// TIA Portal project "FORMING_1500_PLC" (V15)

(* hardware
DEVICE "1.Forming_Machine_PN"  KTP1200 Basic PN
   slot 0: "1.Forming_Machine_PN"  KTP1200 Basic PN  6AV2 123-2MB03-0AX0  15.0.0.0
   slot 1: "HMI_RT_1"  KTP1200 Basic PN  6AV2 123-2MB03-0AX0  15.0.0.0
   slot 5: "Forming_Machine.IE_CP_1"  PROFINET Interface  15.0.0.0
      slot 1: "PROFINET Interface_1"  PROFINET Interface
         slot 1: "Port_1"  Port
DEVICE "GSD device_2"  GSD.Device
   slot 0: "Rack_0"  Rail
DEVICE "GSD device_8"  GSD.Device
   slot 0: "Rack_0"  Rail
DEVICE "GSD device_5"  GSD.Device
   slot 0: "Rack_0"  Rail
DEVICE "GSD device_6"  GSD.Device
   slot 0: "Rack_0"  Rail
DEVICE "GSD device_7"  GSD.Device
   slot 0: "Rack_0"  Rail
DEVICE "GSD device_9"  GSD.Device
   slot 0: "Rack_0"  Rail
DEVICE "GSD device_4"  GSD.Device
   slot 0: "Rack_0"  Rail
DEVICE "GSD device_3"  GSD.Device
   slot 0: "Rack_0"  Rail
DEVICE "GSD device_11"  GSD.Device
   slot 0: "Rack_0"  Rail
DEVICE "GSD device_12"  GSD.Device
   slot 0: "Rack_0"  Rail
DEVICE "GSD device_13"  GSD.Device
   slot 0: "Rack_0"  Rail
DEVICE "GSD device_14"  GSD.Device
   slot 0: "Rack_0"  Rail
DEVICE "GSD device_10"  GSD.Device
   slot 0: "Rack_0"  Rail
DEVICE "GSD device_16"  GSD.Device
   slot 0: "Rack_0"  Rail
DEVICE "GSD device_17"  GSD.Device
   slot 0: "Rack_0"  Rail
DEVICE "GSD device_18"  GSD.Device
   slot 0: "Rack_0"  Rail
DEVICE "GSD device_19"  GSD.Device
   slot 0: "Rack_0"  Rail
DEVICE "GSD device_20"  GSD.Device
   slot 0: "Rack_0"  Rail
DEVICE "GSD device_15"  GSD.Device
   slot 0: "Rack_0"  Rail
DEVICE "GSD device_21"  GSD.Device
   slot 0: "Rack_0"  Rail
DEVICE "GSD device_22"  GSD.Device
   slot 0: "Rack_0"  Rail
DEVICE "GSD device_23"  GSD.Device
   slot 0: "Rack_0"  Rail
DEVICE "S71500/ET200MP station_2"  S7-1500 station
   slot 0: "Rail_0"  Rack  6ES7 590-1***0-0AA0
   slot 0: "PM 190W 120/230VAC"  PM 190W 120/230VAC  6EP1333-4BA00
   slot 1: "FORMING LINE 7 PLC_1"  CPU 1511-1 PN  6ES7 511-1AK02-0AB0  V2.5
      slot 3: "CPU display_1"  6ES7591-1AA00-0AA0
   slot 2: "CM 1542-5_1"  CM 1542-5  6GK7 542-5DX00-0XE0  V2.0
   slot 3: "DI 32x24VDC BA_3"  DI 32x24VDC BA  6ES7 521-1BL10-0AA0  V1.0
   slot 4: "DQ 16x24VDC/0.5A BA_1"  DQ 16x24VDC/0.5A BA  6ES7 522-1BH10-0AA0  V1.0
   slot 5: "DI 32x24VDC BA_1"  DI 32x24VDC BA  6ES7 521-1BL10-0AA0  V1.0
   slot 6: "DI 32x24VDC BA_2"  DI 32x24VDC BA  6ES7 521-1BL10-0AA0  V1.0
*)

// ===== PLC "FORMING LINE 7 PLC_1"  CPU 1511-1 PN =====

VAR_GLOBAL   // PLC tag table "Default tag table"
   "PHOTOCELL OF KIBBLER" AT %I7.4 : Bool;
   "KIBBLER 1 CMD" AT %M28.0 : Bool;
   "KIBBLER CLCKWISE / ANTI CLCKWISE 2" AT %Q124.2 : Bool;
   "KIBBLER 2 CMD" AT %M28.1 : Bool;
   "DELAY KIBBLER 1" AT %T14 : Timer;
   "KIBBLER CLCKWISE / ANTI CLCKWISE 1" AT %Q124.1 : Bool;
   "DELAY KIBBLER 1 RESET" AT %T15 : Timer;
   "DELAY KIBBLER 2" AT %T16 : Timer;
   "DELAY KIBBLER 2 RESET" AT %T17 : Timer;
   "INPUT METAL DETECT ALARM" AT %I7.5 : Bool;
   "input metal detect cmd a" AT %M60.1 : Bool;
   "TIMER RESET ALARM OUT METAL DETECT" AT %T9 : Timer;
   "TIMER INPUT METAL DETECT ALARM" AT %T25 : Timer;
   "input metal detect cmd b" AT %M60.0 : Bool;
   "trigger_alarm_metal_detect" AT %M38.3 : Bool;
   "ALARM OUTPUT WHEN METAL DETECT" AT %Q124.4 : Bool;
   "trigger_time_lap_metal_detect" AT %M38.4 : Bool;
   "TIME LAP WHEN METAL DETECTED" AT %Q124.0 : Bool;
   "RESET TIME LAP WHEN METAL DETECT" AT %T23 : Timer;
   "trigger_sync_addres_13" AT %M31.6 : Bool;
   "trigger_sync_addres_17 a" AT %M32.2 : Bool;
   "trigger_sync_addres_3" AT %M30.4 : Bool;
   "trigger_sync_addres_4" AT %M30.5 : Bool;
   "trigger_sync_addres_5" AT %M30.6 : Bool;
   "trigger_sync_addres_6" AT %M30.7 : Bool;
   "trigger_sync_addres_7" AT %M31.0 : Bool;
   "trigger_sync_addres_8" AT %M31.1 : Bool;
   "trigger_sync_addres_9" AT %M31.2 : Bool;
   "trigger_sync_addres_10" AT %M31.3 : Bool;
   "trigger_sync_addres_11" AT %M31.4 : Bool;
   "trigger_sync_addres_12" AT %M31.5 : Bool;
   "trigger_sync_addres_14" AT %M31.7 : Bool;
   "trigger_sync_addres_15" AT %M32.0 : Bool;
   "trigger_sync_addres_16" AT %M32.1 : Bool;
   "trigger_sync_addres_17 b" AT %M33.2 : Bool;
   "trigger_sync_addres_19" AT %M32.4 : Bool;
   "trigger_sync_addres_21" AT %M32.6 : Bool;
   "trigger_sync_addres_22" AT %M32.7 : Bool;
   "trigger_sync_addres_23" AT %M33.0 : Bool;
   "SB1" AT %I125.0 : Bool;
   "SB2" AT %I125.1 : Bool;
   "SB3" AT %I125.2 : Bool;
   "SB4" AT %I125.3 : Bool;
   "SB5" AT %I125.4 : Bool;
   "SB6" AT %I125.5 : Bool;
   "SB7" AT %I125.6 : Bool;
   "SB8" AT %I125.7 : Bool;
   "SB9" AT %I6.0 : Bool;
   "SB10" AT %I6.1 : Bool;
   "SB11" AT %I6.2 : Bool;
   "SB12" AT %I6.3 : Bool;
   "SB13" AT %I6.4 : Bool;
   "profibus addres 2 fault" AT %M90.1 : Bool;
   "profibus addres 3 fault" AT %M90.2 : Bool;
   "profibus addres 4 fault" AT %M90.3 : Bool;
   "profibus addres 5 fault" AT %M90.4 : Bool;
   "profibus addres 6 fault" AT %M90.5 : Bool;
   "profibus addres 7 fault" AT %M90.6 : Bool;
   "profibus addres 8 fault" AT %M90.7 : Bool;
   "profibus addres 9 fault" AT %M91.0 : Bool;
   "profibus addres 10 fault" AT %M91.1 : Bool;
   "profibus addres 11 fault" AT %M91.2 : Bool;
   "profibus addres 12 fault" AT %M91.3 : Bool;
   "profibus addres 13 fault" AT %M91.4 : Bool;
   "profibus addres 14 fault" AT %M91.5 : Bool;
   "profibus addres 15 fault" AT %M91.6 : Bool;
   "profibus addres 16 fault" AT %M91.7 : Bool;
   "profibus addres 17 fault" AT %M92.0 : Bool;
   "profibus addres 18 fault" AT %M92.1 : Bool;
   "profibus addres 19 fault" AT %M92.2 : Bool;
   "profibus addres 20 fault" AT %M92.3 : Bool;
   "profibus addres 21 fault" AT %M92.4 : Bool;
   "profibus addres 22 fault" AT %M92.5 : Bool;
   "profibus addres 23 fault" AT %M92.6 : Bool;
   "delay10ms_2" AT %T11 : Timer;
   "delay10ms_1" AT %T10 : Timer;
   "delay10ms_4" AT %T13 : Timer;
   "delay10ms_3" AT %T12 : Timer;
   "ROTARY MOULDER MODE" AT %I7.0 : Bool;
   "ROTARY CUTTER MODE" AT %I7.1 : Bool;
   "EMERGENCY" AT %I7.6 : Bool;
   "EMC PRESSED" AT %M92.7 : Bool;
END_VAR

VAR_GLOBAL   // PLC tag table "STEP7 classic symbols"
   "DECREASE_ADDRS_3" AT %I0.5 : Bool;
   "DECREASE_ADDRS_2" AT %I0.3 : Bool;
   "DECREASE_ADDRS_23" AT %I5.5 : Bool;
   "DECREASE_ADDRS_22" AT %I5.3 : Bool;
   "DECREASE_ADDRS_21" AT %I5.1 : Bool;
   "DECREASE_ADDRS_20" AT %I4.7 : Bool;
   "DECREASE_ADDRS_19" AT %I4.5 : Bool;
   "DECREASE_ADDRS_18" AT %I4.3 : Bool;
   "DECREASE_ADDRS_17" AT %I4.1 : Bool;
   "DECREASE_ADDRS_16" AT %I3.7 : Bool;
   "DECREASE_ADDRS_15" AT %I3.5 : Bool;
   "DECREASE_ADDRS_14" AT %I3.3 : Bool;
   "DECREASE_ADDRS_13" AT %I3.1 : Bool;
   "DECREASE_ADDRS_12" AT %I2.7 : Bool;
   "DECREASE_ADDRS_11" AT %I2.5 : Bool;
   "P_MAV_PROFIBUS_23" AT %IW510 : Word;
   "P_CTW_PROFIBUS_7" AT %QW316 : Word;
   "P_CTW_PROFIBUS_6" AT %QW304 : Word;
   "P_CTW_PROFIBUS_5" AT %QW292 : Word;
   "P_CTW_PROFIBUS_4" AT %QW280 : Word;
   "P_CTW_PROFIBUS_3" AT %QW268 : Word;
   "P_CTW_PROFIBUS_2" AT %QW256 : Word;
   "P_CTW_PROFIBUS_11" AT %QW364 : Word;
   "P_CTW_PROFIBUS_10" AT %QW352 : Word;
   "P_CTW_PROFIBUS_9" AT %QW340 : Word;
   "P_CTW_PROFIBUS_8" AT %QW328 : Word;
   "P_CTW_PROFIBUS_13" AT %QW388 : Word;
   "P_CTW_PROFIBUS_12" AT %QW376 : Word;
   "P_CTW_PROFIBUS_15" AT %QW412 : Word;
   "P_CTW_PROFIBUS_14" AT %QW400 : Word;
   "INCREASE_CMD_7" AT %M10.5 : Bool;
   "INCREASE_CMD_6" AT %M10.4 : Bool;
   "INCREASE_CMD_5" AT %M10.3 : Bool;
   "INCREASE_CMD_4" AT %M10.2 : Bool;
   "INCREASE_CMD_3" AT %M10.1 : Bool;
   "INCREASE_CMD_2" AT %M10.0 : Bool;
   "INCREASE_CMD_23" AT %M12.5 : Bool;
   "INCREASE_CMD_22" AT %M12.4 : Bool;
   "INCREASE_CMD_21" AT %M12.3 : Bool;
   "INCREASE_CMD_20" AT %M12.2 : Bool;
   "INCREASE_CMD_19" AT %M12.1 : Bool;
   "INCREASE_CMD_18" AT %M12.0 : Bool;
   "INCREASE_CMD_17" AT %M11.7 : Bool;
   "INCREASE_CMD_16" AT %M11.6 : Bool;
   "INCREASE_CMD_15" AT %M11.5 : Bool;
   "P_MRV_PROFIBUS_8" AT %QW330 : Word;
   "P_MRV_PROFIBUS_7" AT %QW318 : Word;
   "P_MRV_PROFIBUS_12" AT %QW378 : Word;
   "P_MRV_PROFIBUS_11" AT %QW366 : Word;
   "P_MRV_PROFIBUS_10" AT %QW354 : Word;
   "P_MRV_PROFIBUS_15" AT %QW414 : Word;
   "P_MRV_PROFIBUS_14" AT %QW402 : Word;
   "P_MRV_PROFIBUS_13" AT %QW390 : Word;
   "P_MRV_PROFIBUS_18" AT %QW450 : Word;
   "P_MRV_PROFIBUS_17" AT %QW438 : Word;
   "P_MRV_PROFIBUS_16" AT %QW426 : Word;
   "P_MRV_PROFIBUS_21" AT %QW486 : Word;
   "P_MRV_PROFIBUS_20" AT %QW474 : Word;
   "P_MRV_PROFIBUS_19" AT %QW462 : Word;
   "P_MRV_PROFIBUS_22" AT %QW498 : Word;
   "SYNCRON SWIVEL PANNER" AT %I6.7 : Bool;
   "SYNCRON ROTARY CUTTER" AT %I6.6 : Bool;
   "SYNCRON ROTARY MOULDER" AT %I6.5 : Bool;
   "PULSE_1_10_MS" AT %M100.0 : Bool;
   "PULSE_2_10_MS" AT %M100.1 : Bool;
   "HMI_INC_ADDRS_4" AT %M20.3 : Bool;
   "HMI_INC_ADDRS_3" AT %M20.2 : Bool;
   "HMI_INC_ADDRS_2" AT %M20.1 : Bool;
   "HMI_INC_ADDRS_9" AT %M21.0 : Bool;
   "HMI_INC_ADDRS_8" AT %M20.7 : Bool;
   "HMI_INC_ADDRS_7" AT %M20.6 : Bool;
   "HMI_INC_ADDRS_6" AT %M20.5 : Bool;
   "HMI_INC_ADDRS_5" AT %M20.4 : Bool;
   "HMI_INC_ADDRS_21" AT %M22.4 : Bool;
   "HMI_INC_ADDRS_20" AT %M22.3 : Bool;
   "HMI_INC_ADDRS_19" AT %M22.2 : Bool;
   "HMI_INC_ADDRS_18" AT %M22.1 : Bool;
   "HMI_INC_ADDRS_17" AT %M22.0 : Bool;
   "HMI_INC_ADDRS_16" AT %M21.7 : Bool;
   "HMI_INC_ADDRS_15" AT %M21.6 : Bool;
   "P_MAV_PROFIBUS_10" AT %IW354 : Word;
   "P_MAV_PROFIBUS_9" AT %IW342 : Word;
   "P_MAV_PROFIBUS_8" AT %IW330 : Word;
   "P_MAV_PROFIBUS_13" AT %IW390 : Word;
   "P_MAV_PROFIBUS_12" AT %IW378 : Word;
   "P_MAV_PROFIBUS_11" AT %IW366 : Word;
   "P_MAV_PROFIBUS_16" AT %IW426 : Word;
   "P_MAV_PROFIBUS_15" AT %IW414 : Word;
   "P_MAV_PROFIBUS_14" AT %IW402 : Word;
   "P_MAV_PROFIBUS_21" AT %IW486 : Word;
   "P_MAV_PROFIBUS_20" AT %IW474 : Word;
   "P_MAV_PROFIBUS_19" AT %IW462 : Word;
   "P_MAV_PROFIBUS_18" AT %IW450 : Word;
   "P_MAV_PROFIBUS_17" AT %IW438 : Word;
   "P_MAV_PROFIBUS_22" AT %IW498 : Word;
   "HMI_INC_ADDRS_14" AT %M21.5 : Bool;
   "HMI_INC_ADDRS_13" AT %M21.4 : Bool;
   "HMI_INC_ADDRS_12" AT %M21.3 : Bool;
   "HMI_INC_ADDRS_11" AT %M21.2 : Bool;
   "HMI_INC_ADDRS_23" AT %M22.6 : Bool;
   "HMI_INC_ADDRS_22" AT %M22.5 : Bool;
   "HMI_INC_ADDRS_10" AT %M21.1 : Bool;
   "HMI_DEC_ADDRS_14" AT %M25.5 : Bool;
   "HMI_DEC_ADDRS_13" AT %M25.4 : Bool;
   "HMI_DEC_ADDRS_12" AT %M25.3 : Bool;
   "HMI_DEC_ADDRS_11" AT %M25.2 : Bool;
   "HMI_DEC_ADDRS_10" AT %M25.1 : Bool;
   "HMI_DEC_ADDRS_9" AT %M25.0 : Bool;
   "HMI_DEC_ADDRS_8" AT %M24.7 : Bool;
   "HMI_DEC_ADDRS_7" AT %M24.6 : Bool;
   "P_CTW_PROFIBUS_19" AT %QW460 : Word;
   "P_CTW_PROFIBUS_18" AT %QW448 : Word;
   "P_CTW_PROFIBUS_17" AT %QW436 : Word;
   "P_CTW_PROFIBUS_16" AT %QW424 : Word;
   "P_CTW_PROFIBUS_23" AT %QW508 : Word;
   "P_CTW_PROFIBUS_22" AT %QW496 : Word;
   "P_CTW_PROFIBUS_21" AT %QW484 : Word;
   "P_CTW_PROFIBUS_20" AT %QW472 : Word;
   "P_MRV_PROFIBUS_6" AT %QW306 : Word;
   "P_MRV_PROFIBUS_5" AT %QW294 : Word;
   "P_MRV_PROFIBUS_4" AT %QW282 : Word;
   "P_MRV_PROFIBUS_3" AT %QW270 : Word;
   "P_MRV_PROFIBUS_2" AT %QW258 : Word;
   "P_MRV_PROFIBUS_9" AT %QW342 : Word;
   "INCREASE_CMD_14" AT %M11.4 : Bool;
   "INCREASE_CMD_13" AT %M11.3 : Bool;
   "INCREASE_CMD_12" AT %M11.2 : Bool;
   "INCREASE_CMD_11" AT %M11.1 : Bool;
   "INCREASE_CMD_10" AT %M11.0 : Bool;
   "INCREASE_CMD_9" AT %M10.7 : Bool;
   "DECREASE_CMD_2" AT %M15.1 : Bool;
   "DECREASE_CMD_18" AT %M17.1 : Bool;
   "DECREASE_CMD_17" AT %M17.0 : Bool;
   "DECREASE_CMD_16" AT %M16.7 : Bool;
   "DECREASE_CMD_15" AT %M16.6 : Bool;
   "DECREASE_CMD_14" AT %M16.5 : Bool;
   "DECREASE_CMD_13" AT %M16.4 : Bool;
   "DECREASE_CMD_12" AT %M16.3 : Bool;
   "DECREASE_CMD_11" AT %M16.2 : Bool;
   "INCREASE_ADDRS_5" AT %I1.0 : Bool;
   "INCREASE_ADDRS_23" AT %I5.4 : Bool;
   "INCREASE_ADDRS_22" AT %I5.2 : Bool;
   "INCREASE_ADDRS_21" AT %I5.0 : Bool;
   "INCREASE_ADDRS_20" AT %I4.6 : Bool;
   "INCREASE_ADDRS_19" AT %I4.4 : Bool;
   "INCREASE_ADDRS_18" AT %I4.2 : Bool;
   "INCREASE_ADDRS_17" AT %I4.0 : Bool;
   "DECREASE_ADDRS_10" AT %I2.3 : Bool;
   "DECREASE_ADDRS_9" AT %I2.1 : Bool;
   "DECREASE_ADDRS_8" AT %I1.7 : Bool;
   "DECREASE_ADDRS_7" AT %I1.5 : Bool;
   "DECREASE_ADDRS_6" AT %I1.3 : Bool;
   "DECREASE_ADDRS_5" AT %I1.1 : Bool;
   "DECREASE_ADDRS_4" AT %I0.7 : Bool;
   "P_MAV_PROFIBUS_2" AT %IW258 : Word;
   "P_MAV_PROFIBUS_5" AT %IW294 : Word;
   "P_MAV_PROFIBUS_4" AT %IW282 : Word;
   "P_MAV_PROFIBUS_3" AT %IW270 : Word;
   "P_MAV_PROFIBUS_7" AT %IW318 : Word;
   "P_MAV_PROFIBUS_6" AT %IW306 : Word;
   "DECREASE_CMD_10" AT %M16.1 : Bool;
   "DECREASE_CMD_9" AT %M16.0 : Bool;
   "DECREASE_CMD_8" AT %M15.7 : Bool;
   "DECREASE_CMD_7" AT %M15.6 : Bool;
   "DECREASE_CMD_6" AT %M15.5 : Bool;
   "DECREASE_CMD_5" AT %M15.4 : Bool;
   "DECREASE_CMD_4" AT %M15.3 : Bool;
   "DECREASE_CMD_3" AT %M15.2 : Bool;
   "DECREASE_CMD_23" AT %M17.6 : Bool;
   "DECREASE_CMD_22" AT %M17.5 : Bool;
   "DECREASE_CMD_21" AT %M17.4 : Bool;
   "DECREASE_CMD_20" AT %M17.3 : Bool;
   "DECREASE_CMD_19" AT %M17.2 : Bool;
   "P_MRV_PROFIBUS_23" AT %QW510 : Word;
   "INCREASE_ADDRS_4" AT %I0.6 : Bool;
   "INCREASE_ADDRS_3" AT %I0.4 : Bool;
   "INCREASE_ADDRS_2" AT %I0.2 : Bool;
   "INCREASE_ADDRS_16" AT %I3.6 : Bool;
   "INCREASE_ADDRS_15" AT %I3.4 : Bool;
   "INCREASE_ADDRS_14" AT %I3.2 : Bool;
   "INCREASE_ADDRS_13" AT %I3.0 : Bool;
   "INCREASE_ADDRS_12" AT %I2.6 : Bool;
   "INCREASE_ADDRS_11" AT %I2.4 : Bool;
   "INCREASE_ADDRS_10" AT %I2.2 : Bool;
   "INCREASE_ADDRS_9" AT %I2.0 : Bool;
   "INCREASE_ADDRS_8" AT %I1.6 : Bool;
   "INCREASE_ADDRS_7" AT %I1.4 : Bool;
   "INCREASE_ADDRS_6" AT %I1.2 : Bool;
   "HMI_DEC_ADDRS_6" AT %M24.5 : Bool;
   "HMI_DEC_ADDRS_5" AT %M24.4 : Bool;
   "HMI_DEC_ADDRS_4" AT %M24.3 : Bool;
   "HMI_DEC_ADDRS_3" AT %M24.2 : Bool;
   "HMI_DEC_ADDRS_2" AT %M24.1 : Bool;
   "HMI_DEC_ADDRS_23" AT %M26.6 : Bool;
   "HMI_DEC_ADDRS_22" AT %M26.5 : Bool;
   "HMI_DEC_ADDRS_21" AT %M26.4 : Bool;
   "HMI_DEC_ADDRS_20" AT %M26.3 : Bool;
   "HMI_DEC_ADDRS_19" AT %M26.2 : Bool;
   "HMI_DEC_ADDRS_18" AT %M26.1 : Bool;
   "HMI_DEC_ADDRS_17" AT %M26.0 : Bool;
   "HMI_DEC_ADDRS_16" AT %M25.7 : Bool;
   "HMI_DEC_ADDRS_15" AT %M25.6 : Bool;
   "INCREASE_CMD_8" AT %M10.6 : Bool;
   "statusWord_profiBus_2" AT %EW256 : Word;
   "statusWord_profiBus_3" AT %EW268 : Word;
   "statusWord_profiBus_4" AT %EW280 : Word;
   "statusWord_profiBus_5" AT %EW292 : Word;
   "statusWord_profiBus_6" AT %EW304 : Word;
   "statusWord_profiBus_7" AT %EW316 : Word;
   "statusWord_profiBus_8" AT %EW328 : Word;
   "statusWord_profiBus_9" AT %EW340 : Word;
   "statusWord_profiBus_10" AT %EW352 : Word;
   "statusWord_profiBus_11" AT %EW364 : Word;
   "statusWord_profiBus_12" AT %EW376 : Word;
   "statusWord_profiBus_13" AT %EW388 : Word;
   "statusWord_profiBus_14" AT %EW400 : Word;
   "statusWord_profiBus_15" AT %EW412 : Word;
   "statusWord_profiBus_16" AT %EW424 : Word;
   "statusWord_profiBus_17" AT %EW436 : Word;
   "statusWord_profiBus_18" AT %EW448 : Word;
   "statusWord_profiBus_19" AT %EW460 : Word;
   "statusWord_profiBus_20" AT %EW472 : Word;
   "statusWord_profiBus_21" AT %EW484 : Word;
   "statusWord_profiBus_22" AT %EW496 : Word;
   "statusWord_profiBus_23" AT %EW508 : Word;
   "Tag_23" AT %MW66 : Int;
END_VAR

DATA_BLOCK "DB1"   // DB1
{ S7_Optimized_Access := 'FALSE' }
VERSION : 0.1
   VAR
      STAT0 : Int := 1;
      STAT1 : Int;
      STAT2 : Int := 24;
      STAT3 : Int := 1;
      STAT4 : Int := 48;
      STAT5 : Int := 4136;
      STAT6 : Int;
      STAT7 : Int;
      STAT8 : Int;
      STAT9 : Int;
      STAT10 : Int;
      STAT11 : Int;
      STAT12 : Int;
      STAT13 : Int;
      STAT14 : Int;
      STAT15 : Int;
      STAT16 : Int;
      STAT17 : Int;
      STAT18 : Int;
      STAT19 : Int;
      STAT20 : Int;
   END_VAR
BEGIN
END_DATA_BLOCK

DATA_BLOCK "DB2"   // DB2
{ S7_Optimized_Access := 'FALSE' }
VERSION : 0.1
   VAR
      STAT0 : Real;
      STAT1 : Real;
      STAT2 : Real;
      STAT3 : Real;
      STAT4 : Real;
      STAT5 : Real;
      STAT6 : Real;
      STAT7 : Real;
      STAT8 : Real;
      STAT9 : Real;
      STAT10 : Real;
      STAT11 : Real;
      STAT12 : Real;
      STAT13 : Real;
      STAT14 : Real;
      STAT15 : Real;
      STAT16 : Real;
      STAT17 : Real;
      STAT18 : Real;
      STAT19 : Real;
      STAT20 : Real;
      STAT21 : Real;
      STAT22 : Real;
      STAT23 : Real;
      STAT24 : Real;
      STAT25 : Real;
      STAT26 : Real;
      STAT27 : Real;
      STAT28 : Real;
      STAT29 : Real;
      STAT30 : Real;
      STAT31 : Int;
      STAT32 : Int;
      STAT33 : Int;
      STAT34 : Int;
      STAT35 : Int;
   END_VAR
BEGIN
END_DATA_BLOCK

DATA_BLOCK "DB3"   // DB3
{ S7_Optimized_Access := 'FALSE' }
VERSION : 0.1
   VAR
      STAT0 : DInt;
      STAT1 : DInt;
      STAT2 : DInt;
      STAT3 : DInt;
      STAT4 : DInt;
      STAT5 : DInt;
      STAT6 : DInt;
      STAT7 : DInt;
      STAT8 : DInt;
      STAT9 : DInt;
      STAT10 : DInt;
      STAT11 : DInt := DINT#12147;
      STAT12 : DInt := DINT#14276;
      STAT13 : DInt := DINT#14551;
      STAT14 : DInt;
      STAT15 : DInt := DINT#23004;
      STAT16 : DInt;
      STAT17 : DInt;
      STAT18 : DInt;
      STAT19 : DInt;
      STAT20 : DInt;
      STAT21 : DInt;
      STAT22 : DInt;
      STAT23 : DInt;
      STAT24 : DInt;
      STAT25 : DInt;
      STAT26 : DInt;
      STAT27 : DInt;
      STAT28 : DInt;
      STAT29 : DInt;
      STAT30 : DInt;
      STAT31 : DInt := DINT#16386;
      STAT32 : DInt;
      STAT33 : DInt;
      STAT34 : DInt;
      STAT35 : DInt;
      STAT36 : DInt;
      STAT37 : DInt;
      STAT38 : DInt;
      STAT39 : DInt;
      STAT40 : DInt;
      STAT41 : DInt;
      STAT42 : DInt;
      STAT43 : DInt := DINT#12147;
      STAT44 : DInt;
      STAT45 : DInt;
      STAT46 : DInt;
      STAT47 : DInt;
      STAT48 : DInt;
      STAT49 : DInt;
      STAT50 : DInt := DINT#16386;
      STAT51 : DInt;
      STAT52 : DInt;
      STAT53 : DInt;
      STAT54 : DInt;
      STAT55 : DInt;
      STAT56 : DInt;
      STAT57 : DInt;
      STAT58 : DInt;
      STAT59 : DInt;
      STAT60 : DInt;
      STAT61 : DInt;
   END_VAR
BEGIN
END_DATA_BLOCK

DATA_BLOCK "DB4_SPEED_REF"   // DB4
{ S7_Optimized_Access := 'FALSE' }
VERSION : 0.1
   VAR
      MRV_ADDRES_2 : Int := 16386;
      MRV_ADDRES_3 : Int;
      MRV_ADDRES_4 : Int;
      MRV_ADDRES_5 : Int;
      MRV_ADDRES_6 : Int;
      MRV_ADDRES_7 : Int;
      MRV_ADDRES_8 : Int;
      MRV_ADDRES_9 : Int;
      MRV_ADDRES_10 : Int;
      MRV_ADDRES_11 : Int;
      MRV_ADDRES_12 : Int;
      MRV_ADDRES_13 : Int := 12147;
      MRV_ADDRES_14 : Int;
      MRV_ADDRES_15 : Int;
      MRV_ADDRES_16 : Int;
      MRV_ADDRES_17 : Int;
      MRV_ADDRES_18 : Int;
      MRV_ADDRES_19 : Int;
      MRV_ADDRES_20 : Int := 16386;
      MRV_ADDRES_21 : Int;
      MRV_ADDRES_22 : Int;
      MRV_ADDRES_23 : Int;
      STAT22 : Int;
      STAT23 : Int;
      STAT24 : Int;
      STAT25 : Int;
      STAT26 : Int;
      STAT27 : Int;
      STAT28 : Int;
      STAT29 : Int;
      STAT30 : Int;
      STAT31 : Int;
      STAT32 : Int;
      STAT33 : Int;
   END_VAR
BEGIN
END_DATA_BLOCK

DATA_BLOCK "DB5_MAV"   // DB5
{ S7_Optimized_Access := 'FALSE' }
VERSION : 0.1
   VAR
      ADDRES_2 : Int;
      ADDRES_3 : Int;
      ADDRES_4 : Int;
      ADDRES_5 : Int;
      ADDRES_6 : Int;
      ADDRES_7 : Int;
      ADDRES_8 : Int;
      ADDRES_9 : Int;
      ADDRES_10 : Int;
      ADDRES_11 : Int;
      ADDRES_12 : Int;
      ADDRES_13 : Int;
      ADDRES_14 : Int;
      ADDRES_15 : Int;
      ADDRES_16 : Int;
      ADDRES_17 : Int;
      ADDRES_18 : Int;
      ADDRES_19 : Int;
      ADDRES_20 : Int;
      ADDRES_21 : Int;
      ADDRES_22 : Int;
      ADDRES_23 : Int;
      STAT22 : Int;
      STAT23 : Int;
      STAT24 : Int;
      STAT25 : Int;
      STAT26 : Int;
      STAT27 : Int;
      STAT28 : Int;
      STAT29 : Int;
      STAT30 : Int;
      STAT31 : Int;
      STAT32 : Int;
      STAT33 : Int;
      STAT34 : Int;
      STAT35 : Int;
      STAT36 : Int;
      STAT37 : Int;
      STAT38 : Int;
      STAT39 : Int;
   END_VAR
BEGIN
END_DATA_BLOCK

DATA_BLOCK "DB6_MAV2_DBD"   // DB6
{ S7_Optimized_Access := 'FALSE' }
VERSION : 0.1
   VAR
      ADDRES_2 : Real;
      ADDRES_3 : Real;
      ADDRES_4 : Real;
      ADDRES_5 : Real;
      ADDRES_6 : Real;
      ADDRES_7 : Real;
      ADDRES_8 : Real;
      ADDRES_9 : Real;
      ADDRES_10 : Real;
      ADDRES_11 : Real;
      ADDRES_12 : Real;
      ADDRES_13 : Real;
      ADDRES_14 : Real;
      ADDRES_15 : Real;
      ADDRES_16 : Real;
      ADDRES_17 : Real;
      ADDRES_18 : Real;
      ADDRES_19 : Real;
      ADDRES_20 : Real;
      ADDRES_21 : Real;
      ADDRES_22 : Real;
      ADDRES_23 : Real;
      STAT22 : Real;
      STAT23 : Real;
      STAT24 : Real;
      STAT25 : Real;
      STAT26 : Real;
      STAT27 : Real;
      STAT28 : Real;
      SCALLING_2 : Real;
      SCALLING_3 : Real;
      SCALLING_4 : Real;
      SCALLING_5 : Real;
      SCALLING_6 : Real;
      SCALLING_7 : Real;
      SCALLING_8 : Real;
      SCALLING_9 : Real;
      SCALLING_10 : Real;
      SCALLING_11 : Real;
      SCALLING_12 : Real;
      SCALLING_13 : Real;
      SCALLING_14 : Real;
      SCALLING_15 : Real;
      SCALLING_16 : Real;
      SCALLING_17 : Real;
      SCALLING_18 : Real;
      SCALLING_19 : Real;
      SCALLING_20 : Real;
      SCALLING_21 : Real;
      SCALLING_22 : Real;
      SCALLING_23 : Real;
      STAT51 : Real;
      STAT52 : Real;
      STAT53 : Real;
      STAT54 : Real;
      STAT55 : Real;
      STAT56 : Real;
      STAT57 : Real;
      STAT58 : DInt;
      STAT59 : DInt;
      STAT60 : DInt;
      STAT61 : DInt;
      STAT62 : DInt;
      STAT63 : DInt;
      STAT64 : DInt;
      STAT65 : DInt;
      STAT66 : DInt;
      STAT67 : DInt;
      STAT68 : DInt;
      STAT69 : DInt;
      STAT70 : DInt;
      STAT71 : DInt;
      STAT72 : DInt;
      STAT73 : DInt;
      STAT74 : DInt;
      STAT75 : DInt;
      STAT76 : DInt;
      STAT77 : DInt;
      STAT78 : DInt;
      STAT79 : DInt;
      STAT80 : DInt;
      STAT81 : DInt;
      STAT82 : DInt;
      STAT83 : DInt;
      STAT84 : DInt;
      STAT85 : DInt;
      STAT86 : DInt;
      STAT87 : Real;
      STAT88 : Real;
      STAT89 : Real;
      STAT90 : Real;
      STAT91 : DInt;
      STAT92 : DInt;
      STAT93 : Real;
      STAT94 : Real;
      STAT95 : DInt;
      STAT96 : DInt;
   END_VAR
BEGIN
END_DATA_BLOCK

DATA_BLOCK "DB7"   // DB7
{ S7_Optimized_Access := 'FALSE' }
VERSION : 0.1
   VAR
      STAT0 : Word;
      STAT1 : Word;
      STAT2 : Word;
      STAT3 : Word;
      STAT4 : Word;
      STAT5 : Word;
      STAT6 : Word;
      STAT7 : Word;
      STAT8 : Word;
      STAT9 : Word;
      STAT10 : Word;
      STAT11 : Word;
      STAT12 : Word;
      STAT13 : Word;
      STAT14 : Word;
      STAT15 : Word;
      STAT16 : Word;
      STAT17 : Word;
      STAT18 : Word;
      STAT19 : Word;
      STAT20 : Word;
      STAT21 : Word;
      STAT22 : Word;
      STAT23 : Word;
      STAT24 : Word;
      STAT25 : Word;
      STAT26 : Word;
      STAT27 : Word;
      STAT28 : Word;
      STAT29 : Word;
      STAT30 : Word;
      STAT31 : Word;
      STAT32 : Word;
   END_VAR
BEGIN
END_DATA_BLOCK

DATA_BLOCK "DB8_SCALLING_MAV"   // DB8
{ S7_Optimized_Access := 'FALSE' }
VERSION : 0.1
   VAR
      ADDRESS_2 : DInt;
      ADDRESS_3 : DInt;
      ADDRESS_4 : DInt;
      ADDRESS_5 : DInt;
      ADDRESS_6 : DInt;
      ADDRESS_7 : DInt;
      ADDRESS_8 : DInt;
      ADDRESS_9 : DInt;
      ADDRESS_10 : DInt;
      ADDRESS_11 : DInt;
      ADDRESS_12 : DInt;
      ADDRESS_13 : DInt;
      ADDRESS_14 : DInt;
      ADDRESS_15 : DInt;
      ADDRESS_16 : DInt;
      ADDRESS_17 : DInt;
      ADDRESS_18 : DInt;
      ADDRESS_19 : DInt;
      ADDRESS_20 : DInt;
      ADDRESS_21 : DInt;
      ADDRESS_22 : DInt;
      ADDRESS_23 : DInt;
      STAT22 : DInt;
      STAT23 : DInt;
      STAT24 : DInt;
      STAT25 : DInt;
      STAT26 : DInt;
      STAT27 : DInt;
      STAT28 : DInt;
      STAT29 : DInt;
      STAT30 : DInt;
   END_VAR
BEGIN
END_DATA_BLOCK

DATA_BLOCK "DB9"   // DB9
{ S7_Optimized_Access := 'FALSE' }
VERSION : 0.1
   VAR
      STAT0 : Int;
      STAT1 : Int;
   END_VAR
BEGIN
END_DATA_BLOCK

DATA_BLOCK "DB11_RATIO_SYNC"   // DB11
{ S7_Optimized_Access := 'FALSE' }
VERSION : 0.1
   VAR
      STAT0 : Real;
      STAT1 : Real;
      ADDRESS_3 : Real;
      ADDRESS_4 : Real;
      ADDRESS_5 : Real;
      ADDRESS_6 : Real;
      ADDRESS_7 : Real;
      ADDRESS_8 : Real;
      ADDRESS_9 : Real;
      ADDRESS_10 : Real;
      ADDRESS_11 : Real;
      ADDRESS_12 : Real;
      ADDRESS_13 : Real;
      ADDRESS_14 : Real;
      ADDRESS_15 : Real;
      ADDRESS_16 : Real;
      ADDRESS_17 : Real;
      ADDRESS_18 : Real;
      ADDRESS_19 : Real;
      ADDRESS_20 : Real;
      ADDRESS_21 : Real;
      ADDRESS_22 : Real;
      ADDRESS_23 : Real;
      STAT23 : Real;
      STAT24 : Real;
      STAT25 : Real;
      STAT26 : Real;
      STAT27 : Real;
      STAT28 : Real;
      STAT29 : Real;
      STAT30 : Real;
      STAT31 : Real;
      STAT32 : Real;
      STAT33 : Real;
      STAT34 : Real;
      STAT35 : Real;
   END_VAR
BEGIN
END_DATA_BLOCK

DATA_BLOCK "DB12_SPEED_SYNC"   // DB12
{ S7_Optimized_Access := 'FALSE' }
VERSION : 0.1
   VAR
      STAT0 : Real;
      ADDRESS_3 : Real;
      ADDRESS_4 : Real;
      ADDRESS_5 : Real;
      ADDRESS_6 : Real;
      ADDRESS_7 : Real;
      ADDRESS_8 : Real;
      ADDRESS_9 : Real;
      ADDRESS_10 : Real;
      ADDRESS_11 : Real;
      ADDRESS_12 : Real;
      ADDRESS_13 : Real;
      ADDRESS_14 : Real;
      ADDRESS_15 : Real;
      ADDRESS_16 : Real;
      ADDRESS_17 : Real;
      ADDRESS_18 : Real;
      ADDRESS_19 : Real;
      ADDRESS_20 : Real;
      ADDRESS_21 : Real;
      ADDRESS_22 : Real;
      ADDRESS_23 : Real;
      STAT22 : Real;
      STAT23 : Real;
      STAT24 : Real;
      STAT25 : Real;
      STAT26 : Real;
      STAT27 : Real;
      STAT28 : Real;
      STAT29 : Real;
      STAT30 : Real;
      STAT31 : Real;
   END_VAR
BEGIN
END_DATA_BLOCK

DATA_BLOCK "DB13_SPEED_SINGLE_SYNC"   // DB13
{ S7_Optimized_Access := 'FALSE' }
VERSION : 0.1
   VAR
      STAT0 : Real;
      STAT1 : Real;
      ADDRESS_2 : Real := 16386.0;
      ADDRESS_3 : Real;
      ADDRESS_4 : Real;
      ADDRESS_5 : Real;
      ADDRESS_6 : Real;
      ADDRESS_7 : Real;
      ADDRESS_8 : Real;
      ADDRESS_9 : Real;
      ADDRESS_10 : Real;
      ADDRESS_11 : Real;
      ADDRESS_12 : Real;
      ADDRESS_13 : Real;
      ADDRESS_14 : Real;
      ADDRESS_15 : Real;
      ADDRESS_16 : Real;
      ADDRESS_17 : Real;
      ADDRESS_18 : Real;
      ADDRESS_19 : Real;
      ADDRESS_20 : Real := 16386.0;
      ADDRESS_21 : Real;
      ADDRESS_22 : Real;
      ADDRESS_23 : Real;
      STAT24 : Real;
      STAT25 : Real;
      STAT26 : Real;
      STAT27 : Real;
      STAT28 : Real;
      STAT29 : Real;
      STAT30 : Real;
      STAT31 : Real;
      STAT32 : Real;
      STAT33 : Real;
      STAT34 : Real;
   END_VAR
BEGIN
END_DATA_BLOCK

DATA_BLOCK "DB14"   // DB14
{ S7_Optimized_Access := 'FALSE' }
VERSION : 0.1
   VAR
      STAT0 : Word;
      STAT1 : Word;
      STAT2 : Int;
      STAT3 : Word;
      STAT4 : Word;
      STAT5 : Word;
      STAT6 : Bool;
   END_VAR
BEGIN
END_DATA_BLOCK

DATA_BLOCK "DB15_ALARM"   // DB15
{ S7_Optimized_Access := 'FALSE' }
AUTHOR : S4P70
VERSION : 0.1
   VAR
      ALARM_ADDRES_2 : Int;
      ALARM_ADDRES_3 : Int;
      ALARM_ADDRES_4 : Int;
      ALARM_ADDRES_5 : Int;
      ALARM_ADDRES_6 : Int;
      ALARM_ADDRES_7 : Int;
      ALARM_ADDRES_8 : Int;
      ALARM_ADDRES_9 : Int;
      ALARM_ADDRES_10 : Int;
      ALARM_ADDRES_11 : Int;
      ALARM_ADDRES_12 : Int;
      ALARM_ADDRES_13 : Int;
      ALARM_ADDRES_14 : Int;
      ALARM_ADDRES_15 : Int;
      ALARM_ADDRES_16 : Int;
      ALARM_ADDRES_17 : Int;
      ALARM_ADDRES_18 : Int;
      ALARM_ADDRES_19 : Int;
      ALARM_ADDRES_20 : Int;
      ALARM_ADDRES_21 : Int;
      ALARM_ADDRES_22 : Int;
      ALARM_ADDRES_23 : Int;
   END_VAR
BEGIN
END_DATA_BLOCK

DATA_BLOCK "DB16_deviceStates"   // DB16
TITLE = Detect Profibus system
{ S7_Optimized_Access := 'FALSE' }
AUTHOR : sapto
VERSION : 0.1
   VAR
      isLADDR : Hw_IoSystem := 260;
      isMode : UInt := 2;
      returnValue : Int;
      isState : Array[0..1023] of Bool;
   END_VAR
BEGIN
END_DATA_BLOCK

FUNCTION "FC1_KIBBLER & METAL DETECTR" : Void   // FC1, LAD
TITLE = OKIBBLER & METAL DETECTOR
{ S7_Optimized_Access := 'FALSE' }
VERSION : 0.1
   VAR_TEMP   // added for the SCL form of the ladder/FBD networks
      _w1 : Bool;
      _s5time1 : S5Time;
   END_VAR
BEGIN

REGION Network 1: Q124.1 ON SELAMA 15 DETIK SETELAH I7.0 ON SELAMA 5 DETIK
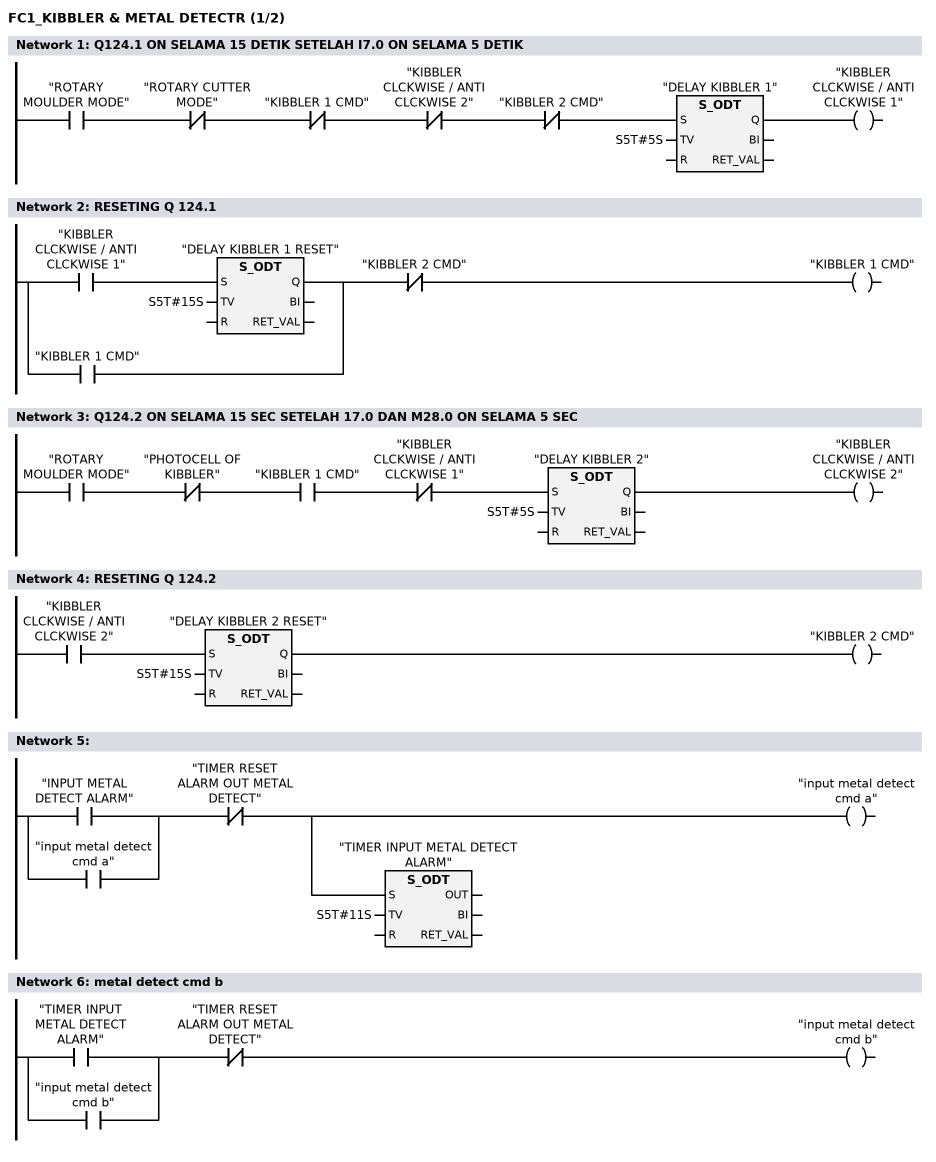
   RUNG wire#powerrail
      Contact( "ROTARY MOULDER MODE" )
      I_Contact( "ROTARY CUTTER MODE" )
      I_Contact( "KIBBLER 1 CMD" )
      I_Contact( "KIBBLER CLCKWISE / ANTI CLCKWISE 2" )
      I_Contact( "KIBBLER 2 CMD" )
      S_ODT(T_NO := "DELAY KIBBLER 1", TV := S5T#5S, R :=, BI =>, RET_VAL =>)
      Coil( "KIBBLER CLCKWISE / ANTI CLCKWISE 1" )
   END_RUNG
   // the same network as SCL:
   #_s5time1 := S_ODT(T_NO := "DELAY KIBBLER 1",
                      S := "ROTARY MOULDER MODE" AND NOT "ROTARY CUTTER MODE" AND NOT "KIBBLER 1 CMD" AND NOT "KIBBLER CLCKWISE / ANTI CLCKWISE 2" AND NOT "KIBBLER 2 CMD",
                      TV := S5T#5S,
                      Q => #_w1);
   "KIBBLER CLCKWISE / ANTI CLCKWISE 1" := #_w1;
END_REGION

REGION Network 2: RESETING Q 124.1
   RUNG wire#powerrail
      Contact( "KIBBLER CLCKWISE / ANTI CLCKWISE 1" )
      S_ODT(T_NO := "DELAY KIBBLER 1 RESET", TV := S5T#15S, R :=, BI =>, RET_VAL =>)
      wire#w1
      I_Contact( "KIBBLER 2 CMD" )
      Coil( "KIBBLER 1 CMD" )
   END_RUNG
   RUNG wire#powerrail
      Contact( "KIBBLER 1 CMD" )
   END_RUNG wire#w1
   // the same network as SCL:
   #_s5time1 := S_ODT(T_NO := "DELAY KIBBLER 1 RESET",
                      S := "KIBBLER CLCKWISE / ANTI CLCKWISE 1",
                      TV := S5T#15S,
                      Q => #_w1);
   "KIBBLER 1 CMD" := (#_w1 OR "KIBBLER 1 CMD") AND NOT "KIBBLER 2 CMD";
END_REGION

REGION Network 3: Q124.2 ON SELAMA 15 SEC SETELAH 17.0 DAN M28.0 ON SELAMA 5 SEC
   RUNG wire#powerrail
      Contact( "ROTARY MOULDER MODE" )
      I_Contact( "PHOTOCELL OF KIBBLER" )
      Contact( "KIBBLER 1 CMD" )
      I_Contact( "KIBBLER CLCKWISE / ANTI CLCKWISE 1" )
      S_ODT(T_NO := "DELAY KIBBLER 2", TV := S5T#5S, R :=, BI =>, RET_VAL =>)
      Coil( "KIBBLER CLCKWISE / ANTI CLCKWISE 2" )
   END_RUNG
   // the same network as SCL:
   #_s5time1 := S_ODT(T_NO := "DELAY KIBBLER 2",
                      S := "ROTARY MOULDER MODE" AND NOT "PHOTOCELL OF KIBBLER" AND "KIBBLER 1 CMD" AND NOT "KIBBLER CLCKWISE / ANTI CLCKWISE 1",
                      TV := S5T#5S,
                      Q => #_w1);
   "KIBBLER CLCKWISE / ANTI CLCKWISE 2" := #_w1;
END_REGION

REGION Network 4: RESETING Q 124.2
   RUNG wire#powerrail
      Contact( "KIBBLER CLCKWISE / ANTI CLCKWISE 2" )
      S_ODT(T_NO := "DELAY KIBBLER 2 RESET", TV := S5T#15S, R :=, BI =>, RET_VAL =>)
      Coil( "KIBBLER 2 CMD" )
   END_RUNG
   // the same network as SCL:
   #_s5time1 := S_ODT(T_NO := "DELAY KIBBLER 2 RESET",
                      S := "KIBBLER CLCKWISE / ANTI CLCKWISE 2",
                      TV := S5T#15S,
                      Q => #_w1);
   "KIBBLER 2 CMD" := #_w1;
END_REGION

REGION Network 5
   RUNG wire#powerrail
      Contact( "INPUT METAL DETECT ALARM" )
      wire#w1
      I_Contact( "TIMER RESET ALARM OUT METAL DETECT" )
      wire#w2
      Coil( "input metal detect cmd a" )
   END_RUNG
   RUNG wire#powerrail
      Contact( "input metal detect cmd a" )
   END_RUNG wire#w1
   RUNG wire#w2
      S_ODT(T_NO := "TIMER INPUT METAL DETECT ALARM", TV := S5T#11S, R :=, BI =>, RET_VAL =>)
   END_RUNG
   // the same network as SCL:
   "input metal detect cmd a" := ("INPUT METAL DETECT ALARM" OR "input metal detect cmd a") AND NOT "TIMER RESET ALARM OUT METAL DETECT";
   #_s5time1 := S_ODT(T_NO := "TIMER INPUT METAL DETECT ALARM", S := "input metal detect cmd a", TV := S5T#11S);
END_REGION

REGION Network 6: metal detect cmd b
   RUNG wire#powerrail
      Contact( "TIMER INPUT METAL DETECT ALARM" )
      wire#w1
      I_Contact( "TIMER RESET ALARM OUT METAL DETECT" )
      Coil( "input metal detect cmd b" )
   END_RUNG
   RUNG wire#powerrail
      Contact( "input metal detect cmd b" )
   END_RUNG wire#w1
   // the same network as SCL:
   "input metal detect cmd b" := ("TIMER INPUT METAL DETECT ALARM" OR "input metal detect cmd b") AND NOT "TIMER RESET ALARM OUT METAL DETECT";
END_REGION